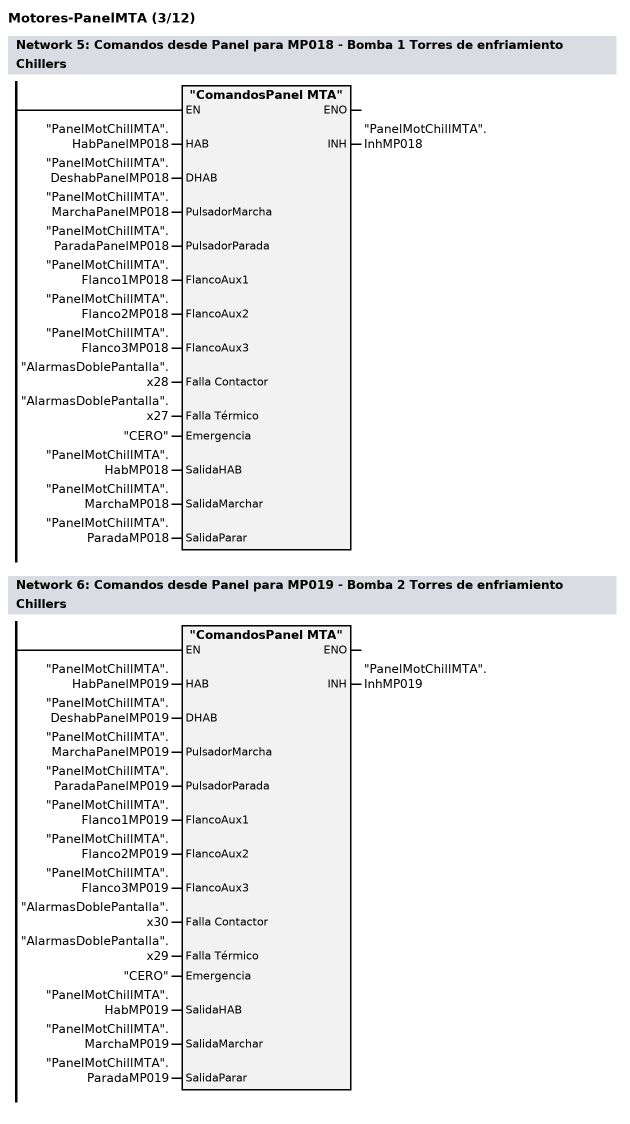
   RUNG wire#powerrail
      "ComandosPanel MTA"(HAB := "PanelMotChillMTA".HabPanelMP018, DHAB := "PanelMotChillMTA".DeshabPanelMP018, PulsadorMarcha := "PanelMotChillMTA".MarchaPanelMP018, PulsadorParada := "PanelMotChillMTA".ParadaPanelMP018, FlancoAux1 := "PanelMotChillMTA".Flanco1MP018, FlancoAux2 := "PanelMotChillMTA".Flanco2MP018, FlancoAux3 := "PanelMotChillMTA".Flanco3MP018, "Falla Contactor" := "AlarmasDoblePantalla".x28, "Falla Térmico" := "AlarmasDoblePantalla".x27, Emergencia := "CERO", SalidaHAB := "PanelMotChillMTA".HabMP018, SalidaMarchar := "PanelMotChillMTA".MarchaMP018, SalidaParar := "PanelMotChillMTA".ParadaMP018, INH => "PanelMotChillMTA".InhMP018)
   END_RUNG
   // the same network as SCL:
   "ComandosPanel MTA"(HAB := "PanelMotChillMTA".HabPanelMP018,
                       DHAB := "PanelMotChillMTA".DeshabPanelMP018,
                       PulsadorMarcha := "PanelMotChillMTA".MarchaPanelMP018,
                       PulsadorParada := "PanelMotChillMTA".ParadaPanelMP018,
                       FlancoAux1 := "PanelMotChillMTA".Flanco1MP018,
                       FlancoAux2 := "PanelMotChillMTA".Flanco2MP018,
                       FlancoAux3 := "PanelMotChillMTA".Flanco3MP018,
                       "Falla Contactor" := "AlarmasDoblePantalla".x28,
                       "Falla Térmico" := "AlarmasDoblePantalla".x27,
                       Emergencia := "CERO",
                       SalidaHAB := "PanelMotChillMTA".HabMP018,
                       SalidaMarchar := "PanelMotChillMTA".MarchaMP018,
                       SalidaParar := "PanelMotChillMTA".ParadaMP018,
                       INH => "PanelMotChillMTA".InhMP018);
END_REGION

REGION Network 6: Comandos desde Panel para MP019 - Bomba 2 Torres de enfriamiento Chillers
   RUNG wire#powerrail
      "ComandosPanel MTA"(HAB := "PanelMotChillMTA".HabPanelMP019, DHAB := "PanelMotChillMTA".DeshabPanelMP019, PulsadorMarcha := "PanelMotChillMTA".MarchaPanelMP019, PulsadorParada := "PanelMotChillMTA".ParadaPanelMP019, FlancoAux1 := "PanelMotChillMTA".Flanco1MP019, FlancoAux2 := "PanelMotChillMTA".Flanco2MP019, FlancoAux3 := "PanelMotChillMTA".Flanco3MP019, "Falla Contactor" := "AlarmasDoblePantalla".x30, "Falla Térmico" := "AlarmasDoblePantalla".x29, Emergencia := "CERO", SalidaHAB := "PanelMotChillMTA".HabMP019, SalidaMarchar := "PanelMotChillMTA".MarchaMP019, SalidaParar := "PanelMotChillMTA".ParadaMP019, INH => "PanelMotChillMTA".InhMP019)
   END_RUNG
   // the same network as SCL:
   "ComandosPanel MTA"(HAB := "PanelMotChillMTA".HabPanelMP019,
                       DHAB := "PanelMotChillMTA".DeshabPanelMP019,
                       PulsadorMarcha := "PanelMotChillMTA".MarchaPanelMP019,
                       PulsadorParada := "PanelMotChillMTA".ParadaPanelMP019,
                       FlancoAux1 := "PanelMotChillMTA".Flanco1MP019,
                       FlancoAux2 := "PanelMotChillMTA".Flanco2MP019,
                       FlancoAux3 := "PanelMotChillMTA".Flanco3MP019,
                       "Falla Contactor" := "AlarmasDoblePantalla".x30,
                       "Falla Térmico" := "AlarmasDoblePantalla".x29,
                       Emergencia := "CERO",
                       SalidaHAB := "PanelMotChillMTA".HabMP019,
                       SalidaMarchar := "PanelMotChillMTA".MarchaMP019,
                       SalidaParar := "PanelMotChillMTA".ParadaMP019,
                       INH => "PanelMotChillMTA".InhMP019);
END_REGION

REGION Network 7: Comandos desde Panel para MT007 - Bomba Soplado L1
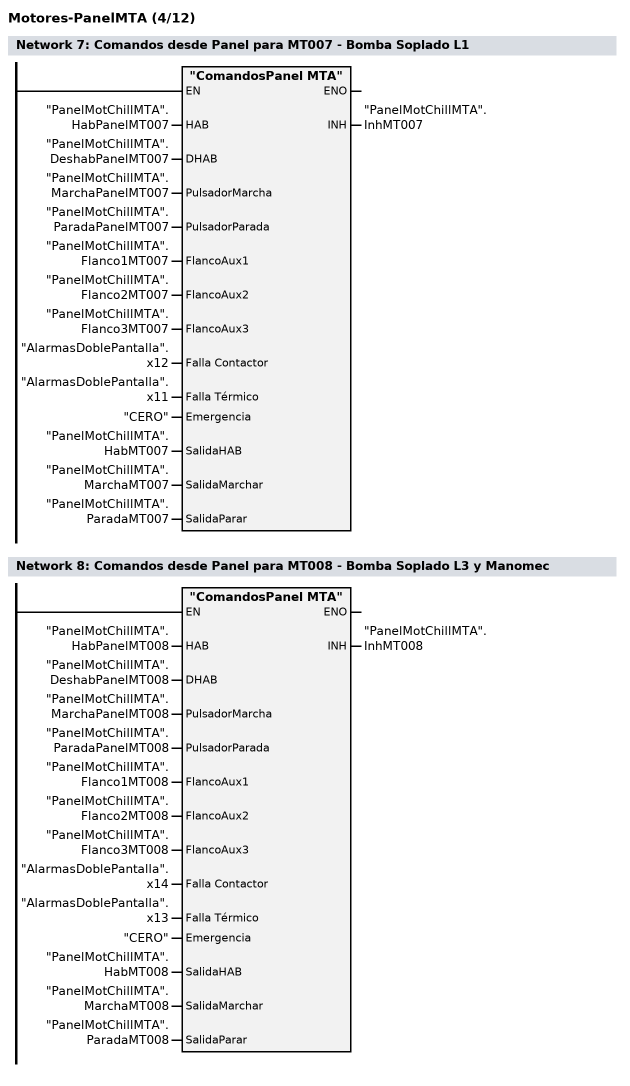
   RUNG wire#powerrail
      "ComandosPanel MTA"(HAB := "PanelMotChillMTA".HabPanelMT007, DHAB := "PanelMotChillMTA".DeshabPanelMT007, PulsadorMarcha := "PanelMotChillMTA".MarchaPanelMT007, PulsadorParada := "PanelMotChillMTA".ParadaPanelMT007, FlancoAux1 := "PanelMotChillMTA".Flanco1MT007, FlancoAux2 := "PanelMotChillMTA".Flanco2MT007, FlancoAux3 := "PanelMotChillMTA".Flanco3MT007, "Falla Contactor" := "AlarmasDoblePantalla".x12, "Falla Térmico" := "AlarmasDoblePantalla".x11, Emergencia := "CERO", INH => "PanelMotChillMTA".InhMT007, SalidaHAB := "PanelMotChillMTA".HabMT007, SalidaMarchar := "PanelMotChillMTA".MarchaMT007, SalidaParar := "PanelMotChillMTA".ParadaMT007)
   END_RUNG
   // the same network as SCL:
   "ComandosPanel MTA"(HAB := "PanelMotChillMTA".HabPanelMT007,
                       DHAB := "PanelMotChillMTA".DeshabPanelMT007,
                       PulsadorMarcha := "PanelMotChillMTA".MarchaPanelMT007,
                       PulsadorParada := "PanelMotChillMTA".ParadaPanelMT007,
                       FlancoAux1 := "PanelMotChillMTA".Flanco1MT007,
                       FlancoAux2 := "PanelMotChillMTA".Flanco2MT007,
                       FlancoAux3 := "PanelMotChillMTA".Flanco3MT007,
                       "Falla Contactor" := "AlarmasDoblePantalla".x12,
                       "Falla Térmico" := "AlarmasDoblePantalla".x11,
                       Emergencia := "CERO",
                       SalidaHAB := "PanelMotChillMTA".HabMT007,
                       SalidaMarchar := "PanelMotChillMTA".MarchaMT007,
                       SalidaParar := "PanelMotChillMTA".ParadaMT007,
                       INH => "PanelMotChillMTA".InhMT007);
END_REGION

REGION Network 8: Comandos desde Panel para MT008 - Bomba Soplado L3 y Manomec
   RUNG wire#powerrail
      "ComandosPanel MTA"(HAB := "PanelMotChillMTA".HabPanelMT008, DHAB := "PanelMotChillMTA".DeshabPanelMT008, PulsadorMarcha := "PanelMotChillMTA".MarchaPanelMT008, PulsadorParada := "PanelMotChillMTA".ParadaPanelMT008, FlancoAux1 := "PanelMotChillMTA".Flanco1MT008, FlancoAux2 := "PanelMotChillMTA".Flanco2MT008, FlancoAux3 := "PanelMotChillMTA".Flanco3MT008, "Falla Contactor" := "AlarmasDoblePantalla".x14, "Falla Térmico" := "AlarmasDoblePantalla".x13, Emergencia := "CERO", INH => "PanelMotChillMTA".InhMT008, SalidaHAB := "PanelMotChillMTA".HabMT008, SalidaMarchar := "PanelMotChillMTA".MarchaMT008, SalidaParar := "PanelMotChillMTA".ParadaMT008)
   END_RUNG
   // the same network as SCL:
   "ComandosPanel MTA"(HAB := "PanelMotChillMTA".HabPanelMT008,
                       DHAB := "PanelMotChillMTA".DeshabPanelMT008,
                       PulsadorMarcha := "PanelMotChillMTA".MarchaPanelMT008,
                       PulsadorParada := "PanelMotChillMTA".ParadaPanelMT008,
                       FlancoAux1 := "PanelMotChillMTA".Flanco1MT008,
                       FlancoAux2 := "PanelMotChillMTA".Flanco2MT008,
                       FlancoAux3 := "PanelMotChillMTA".Flanco3MT008,
                       "Falla Contactor" := "AlarmasDoblePantalla".x14,
                       "Falla Térmico" := "AlarmasDoblePantalla".x13,
                       Emergencia := "CERO",
                       SalidaHAB := "PanelMotChillMTA".HabMT008,
                       SalidaMarchar := "PanelMotChillMTA".MarchaMT008,
                       SalidaParar := "PanelMotChillMTA".ParadaMT008,
                       INH => "PanelMotChillMTA".InhMT008);
END_REGION

REGION Network 9: Comandos desde Panel para MT009 - Bomba Int. L3 y L5
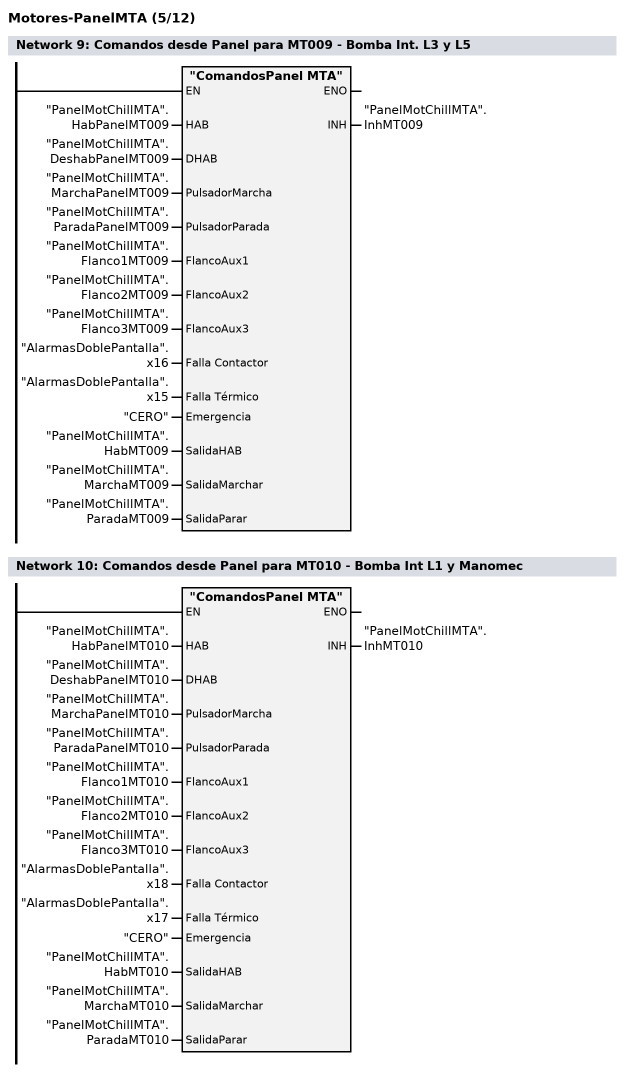
   RUNG wire#powerrail
      "ComandosPanel MTA"(HAB := "PanelMotChillMTA".HabPanelMT009, DHAB := "PanelMotChillMTA".DeshabPanelMT009, PulsadorMarcha := "PanelMotChillMTA".MarchaPanelMT009, PulsadorParada := "PanelMotChillMTA".ParadaPanelMT009, FlancoAux1 := "PanelMotChillMTA".Flanco1MT009, FlancoAux2 := "PanelMotChillMTA".Flanco2MT009, FlancoAux3 := "PanelMotChillMTA".Flanco3MT009, "Falla Contactor" := "AlarmasDoblePantalla".x16, "Falla Térmico" := "AlarmasDoblePantalla".x15, Emergencia := "CERO", INH => "PanelMotChillMTA".InhMT009, SalidaHAB := "PanelMotChillMTA".HabMT009, SalidaMarchar := "PanelMotChillMTA".MarchaMT009, SalidaParar := "PanelMotChillMTA".ParadaMT009)
   END_RUNG
   // the same network as SCL:
   "ComandosPanel MTA"(HAB := "PanelMotChillMTA".HabPanelMT009,
                       DHAB := "PanelMotChillMTA".DeshabPanelMT009,
                       PulsadorMarcha := "PanelMotChillMTA".MarchaPanelMT009,
                       PulsadorParada := "PanelMotChillMTA".ParadaPanelMT009,
                       FlancoAux1 := "PanelMotChillMTA".Flanco1MT009,
                       FlancoAux2 := "PanelMotChillMTA".Flanco2MT009,
                       FlancoAux3 := "PanelMotChillMTA".Flanco3MT009,
                       "Falla Contactor" := "AlarmasDoblePantalla".x16,
                       "Falla Térmico" := "AlarmasDoblePantalla".x15,
                       Emergencia := "CERO",
                       SalidaHAB := "PanelMotChillMTA".HabMT009,
                       SalidaMarchar := "PanelMotChillMTA".MarchaMT009,
                       SalidaParar := "PanelMotChillMTA".ParadaMT009,
                       INH => "PanelMotChillMTA".InhMT009);
END_REGION

REGION Network 10: Comandos desde Panel para MT010 - Bomba Int L1 y Manomec
   RUNG wire#powerrail
      "ComandosPanel MTA"(HAB := "PanelMotChillMTA".HabPanelMT010, DHAB := "PanelMotChillMTA".DeshabPanelMT010, PulsadorMarcha := "PanelMotChillMTA".MarchaPanelMT010, PulsadorParada := "PanelMotChillMTA".ParadaPanelMT010, FlancoAux1 := "PanelMotChillMTA".Flanco1MT010, FlancoAux2 := "PanelMotChillMTA".Flanco2MT010, FlancoAux3 := "PanelMotChillMTA".Flanco3MT010, "Falla Contactor" := "AlarmasDoblePantalla".x18, "Falla Térmico" := "AlarmasDoblePantalla".x17, Emergencia := "CERO", INH => "PanelMotChillMTA".InhMT010, SalidaHAB := "PanelMotChillMTA".HabMT010, SalidaMarchar := "PanelMotChillMTA".MarchaMT010, SalidaParar := "PanelMotChillMTA".ParadaMT010)
   END_RUNG
   // the same network as SCL:
   "ComandosPanel MTA"(HAB := "PanelMotChillMTA".HabPanelMT010,
                       DHAB := "PanelMotChillMTA".DeshabPanelMT010,
                       PulsadorMarcha := "PanelMotChillMTA".MarchaPanelMT010,
                       PulsadorParada := "PanelMotChillMTA".ParadaPanelMT010,
                       FlancoAux1 := "PanelMotChillMTA".Flanco1MT010,
                       FlancoAux2 := "PanelMotChillMTA".Flanco2MT010,
                       FlancoAux3 := "PanelMotChillMTA".Flanco3MT010,
                       "Falla Contactor" := "AlarmasDoblePantalla".x18,
                       "Falla Térmico" := "AlarmasDoblePantalla".x17,
                       Emergencia := "CERO",
                       SalidaHAB := "PanelMotChillMTA".HabMT010,
                       SalidaMarchar := "PanelMotChillMTA".MarchaMT010,
                       SalidaParar := "PanelMotChillMTA".ParadaMT010,
                       INH => "PanelMotChillMTA".InhMT010);
END_REGION

REGION Network 11: Comandos desde Panel para V001 - Ventilador 1 Torres de enfriamiento Chillers
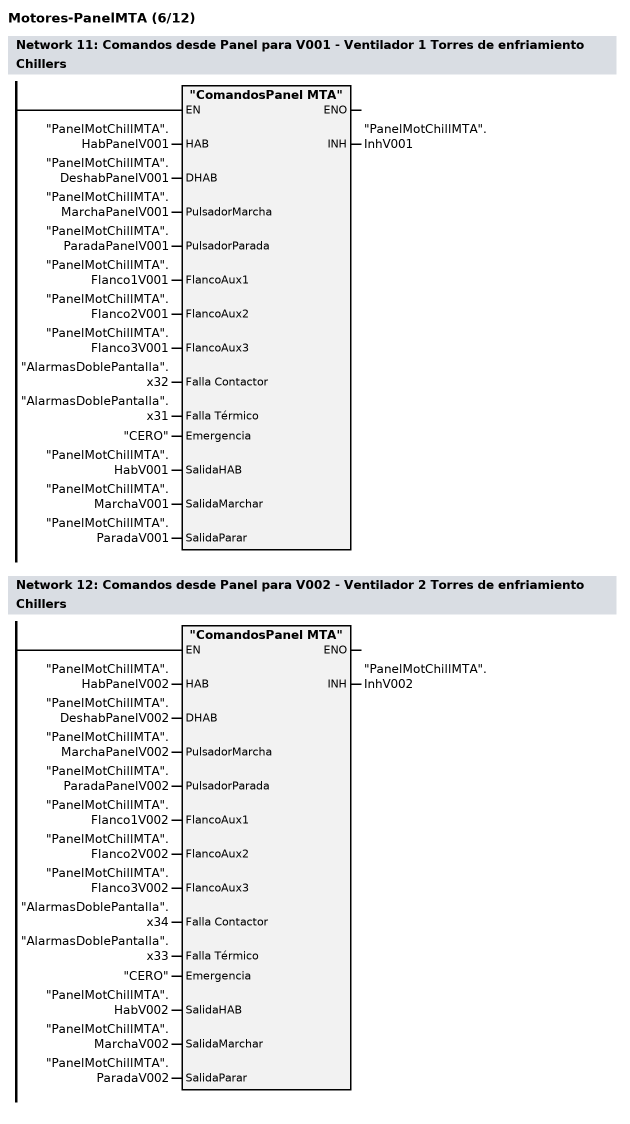
   RUNG wire#powerrail
      "ComandosPanel MTA"(HAB := "PanelMotChillMTA".HabPanelV001, DHAB := "PanelMotChillMTA".DeshabPanelV001, PulsadorMarcha := "PanelMotChillMTA".MarchaPanelV001, PulsadorParada := "PanelMotChillMTA".ParadaPanelV001, FlancoAux1 := "PanelMotChillMTA".Flanco1V001, FlancoAux2 := "PanelMotChillMTA".Flanco2V001, FlancoAux3 := "PanelMotChillMTA".Flanco3V001, "Falla Contactor" := "AlarmasDoblePantalla".x32, "Falla Térmico" := "AlarmasDoblePantalla".x31, Emergencia := "CERO", SalidaHAB := "PanelMotChillMTA".HabV001, SalidaMarchar := "PanelMotChillMTA".MarchaV001, SalidaParar := "PanelMotChillMTA".ParadaV001, INH => "PanelMotChillMTA".InhV001)
   END_RUNG
   // the same network as SCL:
   "ComandosPanel MTA"(HAB := "PanelMotChillMTA".HabPanelV001,
                       DHAB := "PanelMotChillMTA".DeshabPanelV001,
                       PulsadorMarcha := "PanelMotChillMTA".MarchaPanelV001,
                       PulsadorParada := "PanelMotChillMTA".ParadaPanelV001,
                       FlancoAux1 := "PanelMotChillMTA".Flanco1V001,
                       FlancoAux2 := "PanelMotChillMTA".Flanco2V001,
                       FlancoAux3 := "PanelMotChillMTA".Flanco3V001,
                       "Falla Contactor" := "AlarmasDoblePantalla".x32,
                       "Falla Térmico" := "AlarmasDoblePantalla".x31,
                       Emergencia := "CERO",
                       SalidaHAB := "PanelMotChillMTA".HabV001,
                       SalidaMarchar := "PanelMotChillMTA".MarchaV001,
                       SalidaParar := "PanelMotChillMTA".ParadaV001,
                       INH => "PanelMotChillMTA".InhV001);
END_REGION

REGION Network 12: Comandos desde Panel para V002 - Ventilador 2 Torres de enfriamiento Chillers
   RUNG wire#powerrail
      "ComandosPanel MTA"(HAB := "PanelMotChillMTA".HabPanelV002, DHAB := "PanelMotChillMTA".DeshabPanelV002, PulsadorMarcha := "PanelMotChillMTA".MarchaPanelV002, PulsadorParada := "PanelMotChillMTA".ParadaPanelV002, FlancoAux1 := "PanelMotChillMTA".Flanco1V002, FlancoAux2 := "PanelMotChillMTA".Flanco2V002, FlancoAux3 := "PanelMotChillMTA".Flanco3V002, "Falla Contactor" := "AlarmasDoblePantalla".x34, "Falla Térmico" := "AlarmasDoblePantalla".x33, Emergencia := "CERO", SalidaHAB := "PanelMotChillMTA".HabV002, SalidaMarchar := "PanelMotChillMTA".MarchaV002, SalidaParar := "PanelMotChillMTA".ParadaV002, INH => "PanelMotChillMTA".InhV002)
   END_RUNG
   // the same network as SCL:
   "ComandosPanel MTA"(HAB := "PanelMotChillMTA".HabPanelV002,
                       DHAB := "PanelMotChillMTA".DeshabPanelV002,
                       PulsadorMarcha := "PanelMotChillMTA".MarchaPanelV002,
                       PulsadorParada := "PanelMotChillMTA".ParadaPanelV002,
                       FlancoAux1 := "PanelMotChillMTA".Flanco1V002,
                       FlancoAux2 := "PanelMotChillMTA".Flanco2V002,
                       FlancoAux3 := "PanelMotChillMTA".Flanco3V002,
                       "Falla Contactor" := "AlarmasDoblePantalla".x34,
                       "Falla Térmico" := "AlarmasDoblePantalla".x33,
                       Emergencia := "CERO",
                       SalidaHAB := "PanelMotChillMTA".HabV002,
                       SalidaMarchar := "PanelMotChillMTA".MarchaV002,
                       SalidaParar := "PanelMotChillMTA".ParadaV002,
                       INH => "PanelMotChillMTA".InhV002);
END_REGION

REGION Network 13: Comandos desde Panel para V003 - Ventilador 3 Torres de enfriamiento Chillers
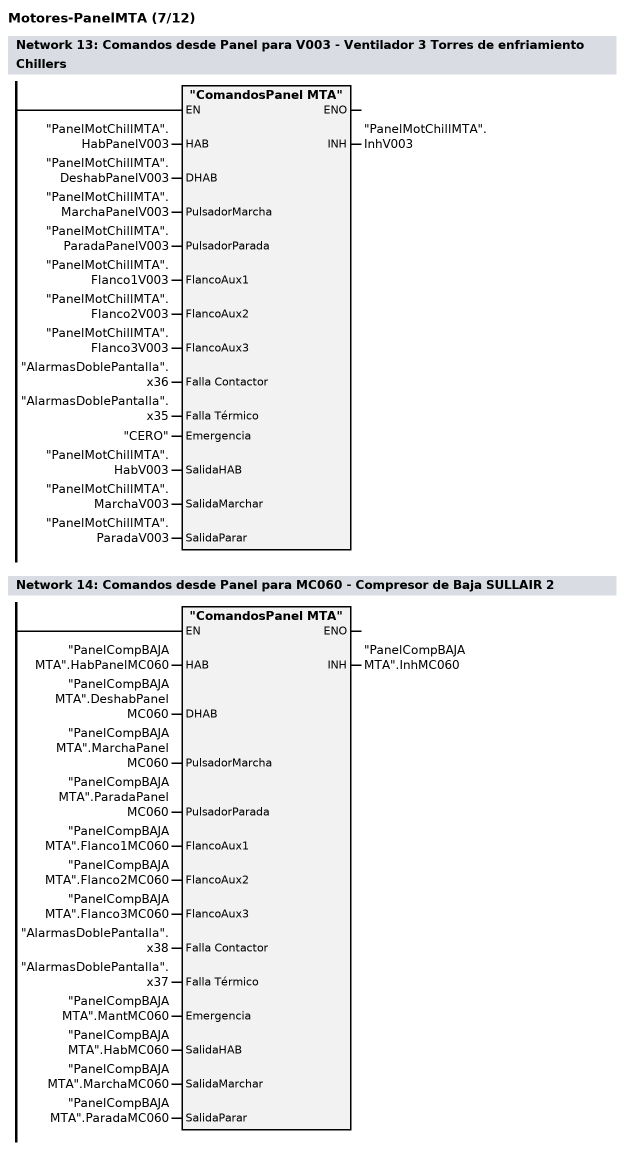
   RUNG wire#powerrail
      "ComandosPanel MTA"(HAB := "PanelMotChillMTA".HabPanelV003, DHAB := "PanelMotChillMTA".DeshabPanelV003, PulsadorMarcha := "PanelMotChillMTA".MarchaPanelV003, PulsadorParada := "PanelMotChillMTA".ParadaPanelV003, FlancoAux1 := "PanelMotChillMTA".Flanco1V003, FlancoAux2 := "PanelMotChillMTA".Flanco2V003, FlancoAux3 := "PanelMotChillMTA".Flanco3V003, "Falla Contactor" := "AlarmasDoblePantalla".x36, "Falla Térmico" := "AlarmasDoblePantalla".x35, Emergencia := "CERO", SalidaHAB := "PanelMotChillMTA".HabV003, SalidaMarchar := "PanelMotChillMTA".MarchaV003, SalidaParar := "PanelMotChillMTA".ParadaV003, INH => "PanelMotChillMTA".InhV003)
   END_RUNG
   // the same network as SCL:
   "ComandosPanel MTA"(HAB := "PanelMotChillMTA".HabPanelV003,
                       DHAB := "PanelMotChillMTA".DeshabPanelV003,
                       PulsadorMarcha := "PanelMotChillMTA".MarchaPanelV003,
                       PulsadorParada := "PanelMotChillMTA".ParadaPanelV003,
                       FlancoAux1 := "PanelMotChillMTA".Flanco1V003,
                       FlancoAux2 := "PanelMotChillMTA".Flanco2V003,
                       FlancoAux3 := "PanelMotChillMTA".Flanco3V003,
                       "Falla Contactor" := "AlarmasDoblePantalla".x36,
                       "Falla Térmico" := "AlarmasDoblePantalla".x35,
                       Emergencia := "CERO",
                       SalidaHAB := "PanelMotChillMTA".HabV003,
                       SalidaMarchar := "PanelMotChillMTA".MarchaV003,
                       SalidaParar := "PanelMotChillMTA".ParadaV003,
                       INH => "PanelMotChillMTA".InhV003);
END_REGION

REGION Network 14: Comandos desde Panel para MC060 - Compresor de Baja SULLAIR 2
   RUNG wire#powerrail
      "ComandosPanel MTA"(HAB := "PanelCompBAJA MTA".HabPanelMC060, DHAB := "PanelCompBAJA MTA".DeshabPanelMC060, PulsadorMarcha := "PanelCompBAJA MTA".MarchaPanelMC060, PulsadorParada := "PanelCompBAJA MTA".ParadaPanelMC060, FlancoAux1 := "PanelCompBAJA MTA".Flanco1MC060, FlancoAux2 := "PanelCompBAJA MTA".Flanco2MC060, FlancoAux3 := "PanelCompBAJA MTA".Flanco3MC060, "Falla Contactor" := "AlarmasDoblePantalla".x38, "Falla Térmico" := "AlarmasDoblePantalla".x37, Emergencia := "PanelCompBAJA MTA".MantMC060, INH => "PanelCompBAJA MTA".InhMC060, SalidaHAB := "PanelCompBAJA MTA".HabMC060, SalidaMarchar := "PanelCompBAJA MTA".MarchaMC060, SalidaParar := "PanelCompBAJA MTA".ParadaMC060)
   END_RUNG
   // the same network as SCL:
   "ComandosPanel MTA"(HAB := "PanelCompBAJA MTA".HabPanelMC060,
                       DHAB := "PanelCompBAJA MTA".DeshabPanelMC060,
                       PulsadorMarcha := "PanelCompBAJA MTA".MarchaPanelMC060,
                       PulsadorParada := "PanelCompBAJA MTA".ParadaPanelMC060,
                       FlancoAux1 := "PanelCompBAJA MTA".Flanco1MC060,
                       FlancoAux2 := "PanelCompBAJA MTA".Flanco2MC060,
                       FlancoAux3 := "PanelCompBAJA MTA".Flanco3MC060,
                       "Falla Contactor" := "AlarmasDoblePantalla".x38,
                       "Falla Térmico" := "AlarmasDoblePantalla".x37,
                       Emergencia := "PanelCompBAJA MTA".MantMC060,
                       SalidaHAB := "PanelCompBAJA MTA".HabMC060,
                       SalidaMarchar := "PanelCompBAJA MTA".MarchaMC060,
                       SalidaParar := "PanelCompBAJA MTA".ParadaMC060,
                       INH => "PanelCompBAJA MTA".InhMC060);
END_REGION

REGION Network 15: Comandos desde Panel para MC061 - Compresor de Baja SULLAIR 1
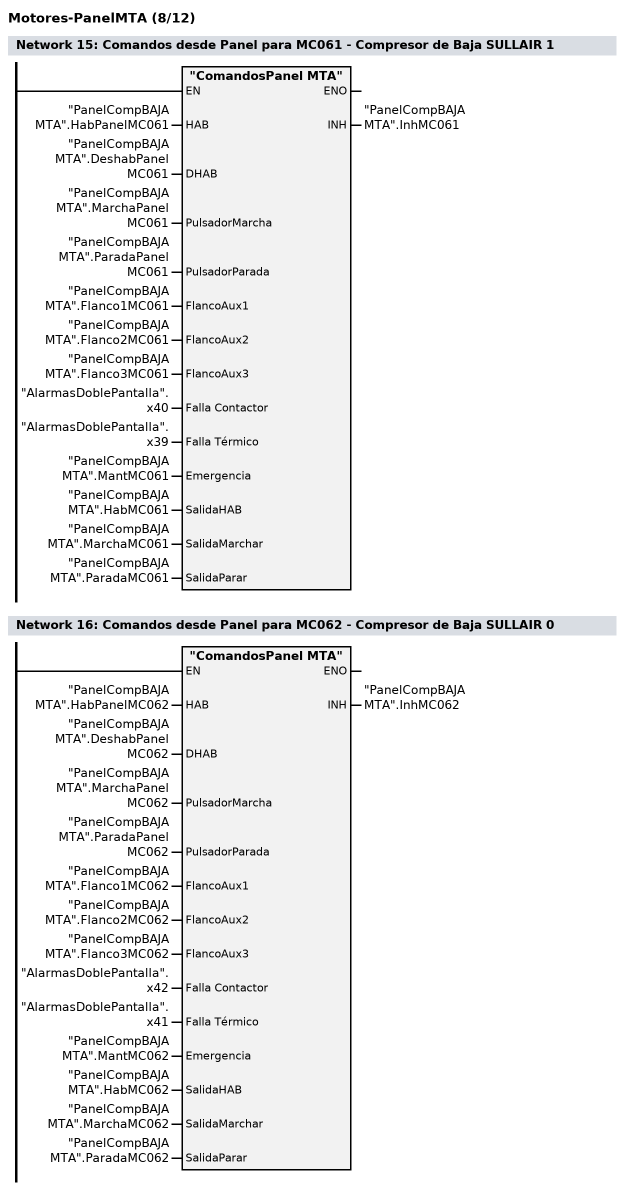
   RUNG wire#powerrail
      "ComandosPanel MTA"(HAB := "PanelCompBAJA MTA".HabPanelMC061, DHAB := "PanelCompBAJA MTA".DeshabPanelMC061, PulsadorMarcha := "PanelCompBAJA MTA".MarchaPanelMC061, PulsadorParada := "PanelCompBAJA MTA".ParadaPanelMC061, FlancoAux1 := "PanelCompBAJA MTA".Flanco1MC061, FlancoAux2 := "PanelCompBAJA MTA".Flanco2MC061, FlancoAux3 := "PanelCompBAJA MTA".Flanco3MC061, "Falla Contactor" := "AlarmasDoblePantalla".x40, "Falla Térmico" := "AlarmasDoblePantalla".x39, Emergencia := "PanelCompBAJA MTA".MantMC061, INH => "PanelCompBAJA MTA".InhMC061, SalidaHAB := "PanelCompBAJA MTA".HabMC061, SalidaMarchar := "PanelCompBAJA MTA".MarchaMC061, SalidaParar := "PanelCompBAJA MTA".ParadaMC061)
   END_RUNG
   // the same network as SCL:
   "ComandosPanel MTA"(HAB := "PanelCompBAJA MTA".HabPanelMC061,
                       DHAB := "PanelCompBAJA MTA".DeshabPanelMC061,
                       PulsadorMarcha := "PanelCompBAJA MTA".MarchaPanelMC061,
                       PulsadorParada := "PanelCompBAJA MTA".ParadaPanelMC061,
                       FlancoAux1 := "PanelCompBAJA MTA".Flanco1MC061,
                       FlancoAux2 := "PanelCompBAJA MTA".Flanco2MC061,
                       FlancoAux3 := "PanelCompBAJA MTA".Flanco3MC061,
                       "Falla Contactor" := "AlarmasDoblePantalla".x40,
                       "Falla Térmico" := "AlarmasDoblePantalla".x39,
                       Emergencia := "PanelCompBAJA MTA".MantMC061,
                       SalidaHAB := "PanelCompBAJA MTA".HabMC061,
                       SalidaMarchar := "PanelCompBAJA MTA".MarchaMC061,
                       SalidaParar := "PanelCompBAJA MTA".ParadaMC061,
                       INH => "PanelCompBAJA MTA".InhMC061);
END_REGION

REGION Network 16: Comandos desde Panel para MC062 - Compresor de Baja SULLAIR 0
   RUNG wire#powerrail
      "ComandosPanel MTA"(HAB := "PanelCompBAJA MTA".HabPanelMC062, DHAB := "PanelCompBAJA MTA".DeshabPanelMC062, PulsadorMarcha := "PanelCompBAJA MTA".MarchaPanelMC062, PulsadorParada := "PanelCompBAJA MTA".ParadaPanelMC062, FlancoAux1 := "PanelCompBAJA MTA".Flanco1MC062, FlancoAux2 := "PanelCompBAJA MTA".Flanco2MC062, FlancoAux3 := "PanelCompBAJA MTA".Flanco3MC062, "Falla Contactor" := "AlarmasDoblePantalla".x42, "Falla Térmico" := "AlarmasDoblePantalla".x41, Emergencia := "PanelCompBAJA MTA".MantMC062, INH => "PanelCompBAJA MTA".InhMC062, SalidaHAB := "PanelCompBAJA MTA".HabMC062, SalidaMarchar := "PanelCompBAJA MTA".MarchaMC062, SalidaParar := "PanelCompBAJA MTA".ParadaMC062)
   END_RUNG
   // the same network as SCL:
   "ComandosPanel MTA"(HAB := "PanelCompBAJA MTA".HabPanelMC062,
                       DHAB := "PanelCompBAJA MTA".DeshabPanelMC062,
                       PulsadorMarcha := "PanelCompBAJA MTA".MarchaPanelMC062,
                       PulsadorParada := "PanelCompBAJA MTA".ParadaPanelMC062,
                       FlancoAux1 := "PanelCompBAJA MTA".Flanco1MC062,
                       FlancoAux2 := "PanelCompBAJA MTA".Flanco2MC062,
                       FlancoAux3 := "PanelCompBAJA MTA".Flanco3MC062,
                       "Falla Contactor" := "AlarmasDoblePantalla".x42,
                       "Falla Térmico" := "AlarmasDoblePantalla".x41,
                       Emergencia := "PanelCompBAJA MTA".MantMC062,
                       SalidaHAB := "PanelCompBAJA MTA".HabMC062,
                       SalidaMarchar := "PanelCompBAJA MTA".MarchaMC062,
                       SalidaParar := "PanelCompBAJA MTA".ParadaMC062,
                       INH => "PanelCompBAJA MTA".InhMC062);
END_REGION

REGION Network 17: Comandos desde Panel para MC063 - Compresor de Baja ATLAS 3
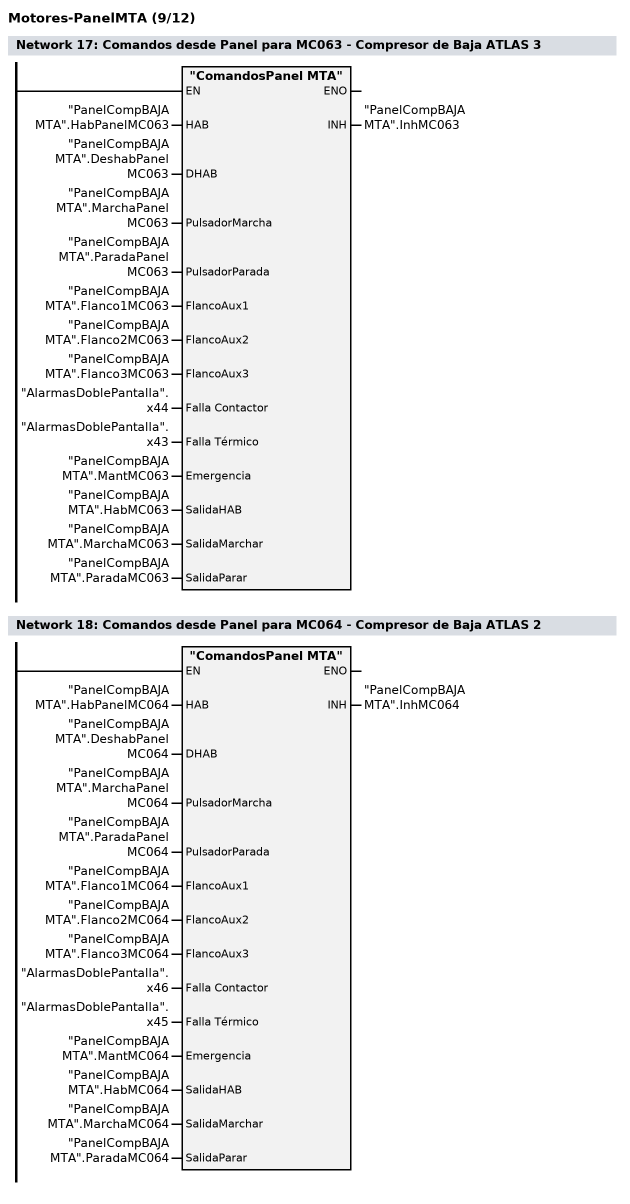
   RUNG wire#powerrail
      "ComandosPanel MTA"(HAB := "PanelCompBAJA MTA".HabPanelMC063, DHAB := "PanelCompBAJA MTA".DeshabPanelMC063, PulsadorMarcha := "PanelCompBAJA MTA".MarchaPanelMC063, PulsadorParada := "PanelCompBAJA MTA".ParadaPanelMC063, FlancoAux1 := "PanelCompBAJA MTA".Flanco1MC063, FlancoAux2 := "PanelCompBAJA MTA".Flanco2MC063, FlancoAux3 := "PanelCompBAJA MTA".Flanco3MC063, "Falla Contactor" := "AlarmasDoblePantalla".x44, "Falla Térmico" := "AlarmasDoblePantalla".x43, Emergencia := "PanelCompBAJA MTA".MantMC063, INH => "PanelCompBAJA MTA".InhMC063, SalidaHAB := "PanelCompBAJA MTA".HabMC063, SalidaMarchar := "PanelCompBAJA MTA".MarchaMC063, SalidaParar := "PanelCompBAJA MTA".ParadaMC063)
   END_RUNG
   // the same network as SCL:
   "ComandosPanel MTA"(HAB := "PanelCompBAJA MTA".HabPanelMC063,
                       DHAB := "PanelCompBAJA MTA".DeshabPanelMC063,
                       PulsadorMarcha := "PanelCompBAJA MTA".MarchaPanelMC063,
                       PulsadorParada := "PanelCompBAJA MTA".ParadaPanelMC063,
                       FlancoAux1 := "PanelCompBAJA MTA".Flanco1MC063,
                       FlancoAux2 := "PanelCompBAJA MTA".Flanco2MC063,
                       FlancoAux3 := "PanelCompBAJA MTA".Flanco3MC063,
                       "Falla Contactor" := "AlarmasDoblePantalla".x44,
                       "Falla Térmico" := "AlarmasDoblePantalla".x43,
                       Emergencia := "PanelCompBAJA MTA".MantMC063,
                       SalidaHAB := "PanelCompBAJA MTA".HabMC063,
                       SalidaMarchar := "PanelCompBAJA MTA".MarchaMC063,
                       SalidaParar := "PanelCompBAJA MTA".ParadaMC063,
                       INH => "PanelCompBAJA MTA".InhMC063);
END_REGION

REGION Network 18: Comandos desde Panel para MC064 - Compresor de Baja ATLAS 2
   RUNG wire#powerrail
      "ComandosPanel MTA"(HAB := "PanelCompBAJA MTA".HabPanelMC064, DHAB := "PanelCompBAJA MTA".DeshabPanelMC064, PulsadorMarcha := "PanelCompBAJA MTA".MarchaPanelMC064, PulsadorParada := "PanelCompBAJA MTA".ParadaPanelMC064, FlancoAux1 := "PanelCompBAJA MTA".Flanco1MC064, FlancoAux2 := "PanelCompBAJA MTA".Flanco2MC064, FlancoAux3 := "PanelCompBAJA MTA".Flanco3MC064, "Falla Contactor" := "AlarmasDoblePantalla".x46, "Falla Térmico" := "AlarmasDoblePantalla".x45, Emergencia := "PanelCompBAJA MTA".MantMC064, INH => "PanelCompBAJA MTA".InhMC064, SalidaHAB := "PanelCompBAJA MTA".HabMC064, SalidaMarchar := "PanelCompBAJA MTA".MarchaMC064, SalidaParar := "PanelCompBAJA MTA".ParadaMC064)
   END_RUNG
   // the same network as SCL:
   "ComandosPanel MTA"(HAB := "PanelCompBAJA MTA".HabPanelMC064,
                       DHAB := "PanelCompBAJA MTA".DeshabPanelMC064,
                       PulsadorMarcha := "PanelCompBAJA MTA".MarchaPanelMC064,
                       PulsadorParada := "PanelCompBAJA MTA".ParadaPanelMC064,
                       FlancoAux1 := "PanelCompBAJA MTA".Flanco1MC064,
                       FlancoAux2 := "PanelCompBAJA MTA".Flanco2MC064,
                       FlancoAux3 := "PanelCompBAJA MTA".Flanco3MC064,
                       "Falla Contactor" := "AlarmasDoblePantalla".x46,
                       "Falla Térmico" := "AlarmasDoblePantalla".x45,
                       Emergencia := "PanelCompBAJA MTA".MantMC064,
                       SalidaHAB := "PanelCompBAJA MTA".HabMC064,
                       SalidaMarchar := "PanelCompBAJA MTA".MarchaMC064,
                       SalidaParar := "PanelCompBAJA MTA".ParadaMC064,
                       INH => "PanelCompBAJA MTA".InhMC064);
END_REGION

REGION Network 19: Comandos desde Panel para MS050 - Secador de Alta ABC1
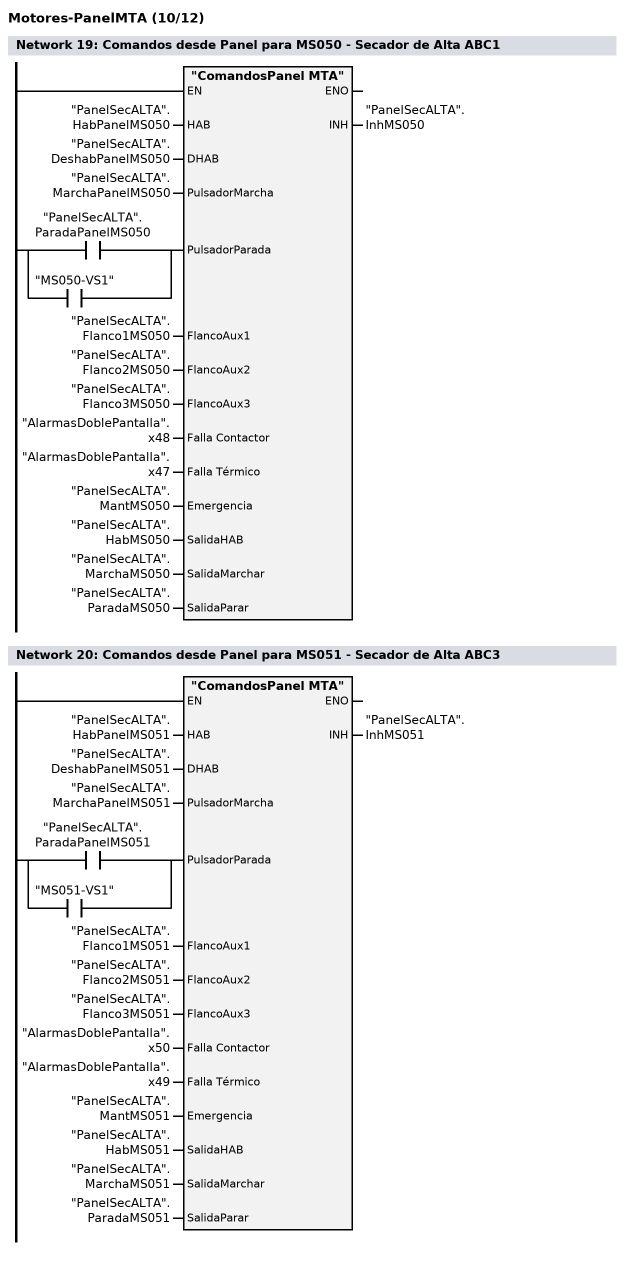
   RUNG wire#powerrail
      "ComandosPanel MTA"(HAB := "PanelSecALTA".HabPanelMS050, DHAB := "PanelSecALTA".DeshabPanelMS050, PulsadorMarcha := "PanelSecALTA".MarchaPanelMS050, PulsadorParada := wire#w1, FlancoAux1 := "PanelSecALTA".Flanco1MS050, FlancoAux2 := "PanelSecALTA".Flanco2MS050, FlancoAux3 := "PanelSecALTA".Flanco3MS050, "Falla Contactor" := "AlarmasDoblePantalla".x48, "Falla Térmico" := "AlarmasDoblePantalla".x47, Emergencia := "PanelSecALTA".MantMS050, INH => "PanelSecALTA".InhMS050, SalidaHAB := "PanelSecALTA".HabMS050, SalidaMarchar := "PanelSecALTA".MarchaMS050, SalidaParar := "PanelSecALTA".ParadaMS050)
   END_RUNG
   RUNG wire#powerrail
      Contact( "PanelSecALTA".ParadaPanelMS050 )
   END_RUNG wire#w1
   RUNG wire#powerrail
      Contact( "MS050-VS1" )
   END_RUNG wire#w1
   // the same network as SCL:
   "ComandosPanel MTA"(HAB := "PanelSecALTA".HabPanelMS050,
                       DHAB := "PanelSecALTA".DeshabPanelMS050,
                       PulsadorMarcha := "PanelSecALTA".MarchaPanelMS050,
                       PulsadorParada := "PanelSecALTA".ParadaPanelMS050 OR "MS050-VS1",
                       FlancoAux1 := "PanelSecALTA".Flanco1MS050,
                       FlancoAux2 := "PanelSecALTA".Flanco2MS050,
                       FlancoAux3 := "PanelSecALTA".Flanco3MS050,
                       "Falla Contactor" := "AlarmasDoblePantalla".x48,
                       "Falla Térmico" := "AlarmasDoblePantalla".x47,
                       Emergencia := "PanelSecALTA".MantMS050,
                       SalidaHAB := "PanelSecALTA".HabMS050,
                       SalidaMarchar := "PanelSecALTA".MarchaMS050,
                       SalidaParar := "PanelSecALTA".ParadaMS050,
                       INH => "PanelSecALTA".InhMS050);
END_REGION

REGION Network 20: Comandos desde Panel para MS051 - Secador de Alta ABC3
   RUNG wire#powerrail
      "ComandosPanel MTA"(HAB := "PanelSecALTA".HabPanelMS051, DHAB := "PanelSecALTA".DeshabPanelMS051, PulsadorMarcha := "PanelSecALTA".MarchaPanelMS051, PulsadorParada := wire#w1, FlancoAux1 := "PanelSecALTA".Flanco1MS051, FlancoAux2 := "PanelSecALTA".Flanco2MS051, FlancoAux3 := "PanelSecALTA".Flanco3MS051, "Falla Contactor" := "AlarmasDoblePantalla".x50, "Falla Térmico" := "AlarmasDoblePantalla".x49, Emergencia := "PanelSecALTA".MantMS051, INH => "PanelSecALTA".InhMS051, SalidaHAB := "PanelSecALTA".HabMS051, SalidaMarchar := "PanelSecALTA".MarchaMS051, SalidaParar := "PanelSecALTA".ParadaMS051)
   END_RUNG
   RUNG wire#powerrail
      Contact( "PanelSecALTA".ParadaPanelMS051 )
   END_RUNG wire#w1
   RUNG wire#powerrail
      Contact( "MS051-VS1" )
   END_RUNG wire#w1
   // the same network as SCL:
   "ComandosPanel MTA"(HAB := "PanelSecALTA".HabPanelMS051,
                       DHAB := "PanelSecALTA".DeshabPanelMS051,
                       PulsadorMarcha := "PanelSecALTA".MarchaPanelMS051,
                       PulsadorParada := "PanelSecALTA".ParadaPanelMS051 OR "MS051-VS1",
                       FlancoAux1 := "PanelSecALTA".Flanco1MS051,
                       FlancoAux2 := "PanelSecALTA".Flanco2MS051,
                       FlancoAux3 := "PanelSecALTA".Flanco3MS051,
                       "Falla Contactor" := "AlarmasDoblePantalla".x50,
                       "Falla Térmico" := "AlarmasDoblePantalla".x49,
                       Emergencia := "PanelSecALTA".MantMS051,
                       SalidaHAB := "PanelSecALTA".HabMS051,
                       SalidaMarchar := "PanelSecALTA".MarchaMS051,
                       SalidaParar := "PanelSecALTA".ParadaMS051,
                       INH => "PanelSecALTA".InhMS051);
END_REGION

REGION Network 21: Comandos desde Panel para MS052 - Secador de Alta ABC2
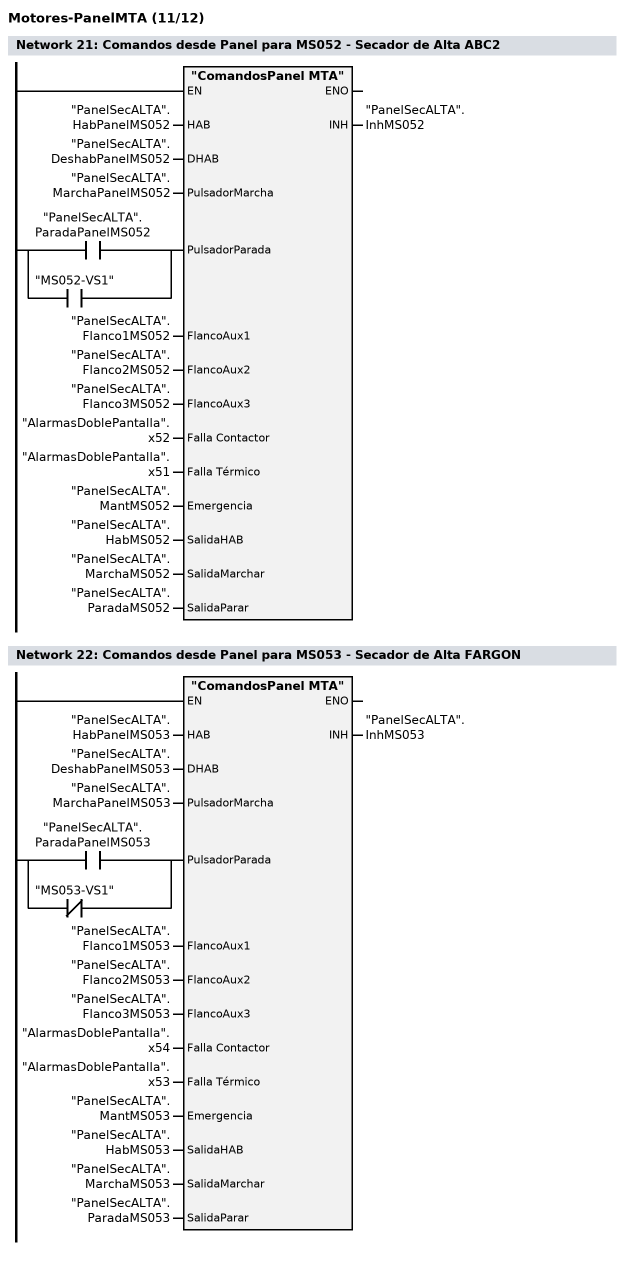
   RUNG wire#powerrail
      "ComandosPanel MTA"(HAB := "PanelSecALTA".HabPanelMS052, DHAB := "PanelSecALTA".DeshabPanelMS052, PulsadorMarcha := "PanelSecALTA".MarchaPanelMS052, PulsadorParada := wire#w1, FlancoAux1 := "PanelSecALTA".Flanco1MS052, FlancoAux2 := "PanelSecALTA".Flanco2MS052, FlancoAux3 := "PanelSecALTA".Flanco3MS052, "Falla Contactor" := "AlarmasDoblePantalla".x52, "Falla Térmico" := "AlarmasDoblePantalla".x51, Emergencia := "PanelSecALTA".MantMS052, INH => "PanelSecALTA".InhMS052, SalidaHAB := "PanelSecALTA".HabMS052, SalidaMarchar := "PanelSecALTA".MarchaMS052, SalidaParar := "PanelSecALTA".ParadaMS052)
   END_RUNG
   RUNG wire#powerrail
      Contact( "PanelSecALTA".ParadaPanelMS052 )
   END_RUNG wire#w1
   RUNG wire#powerrail
      Contact( "MS052-VS1" )
   END_RUNG wire#w1
   // the same network as SCL:
   "ComandosPanel MTA"(HAB := "PanelSecALTA".HabPanelMS052,
                       DHAB := "PanelSecALTA".DeshabPanelMS052,
                       PulsadorMarcha := "PanelSecALTA".MarchaPanelMS052,
                       PulsadorParada := "PanelSecALTA".ParadaPanelMS052 OR "MS052-VS1",
                       FlancoAux1 := "PanelSecALTA".Flanco1MS052,
                       FlancoAux2 := "PanelSecALTA".Flanco2MS052,
                       FlancoAux3 := "PanelSecALTA".Flanco3MS052,
                       "Falla Contactor" := "AlarmasDoblePantalla".x52,
                       "Falla Térmico" := "AlarmasDoblePantalla".x51,
                       Emergencia := "PanelSecALTA".MantMS052,
                       SalidaHAB := "PanelSecALTA".HabMS052,
                       SalidaMarchar := "PanelSecALTA".MarchaMS052,
                       SalidaParar := "PanelSecALTA".ParadaMS052,
                       INH => "PanelSecALTA".InhMS052);
END_REGION

REGION Network 22: Comandos desde Panel para MS053 - Secador de Alta FARGON
   RUNG wire#powerrail
      "ComandosPanel MTA"(HAB := "PanelSecALTA".HabPanelMS053, DHAB := "PanelSecALTA".DeshabPanelMS053, PulsadorMarcha := "PanelSecALTA".MarchaPanelMS053, PulsadorParada := wire#w1, FlancoAux1 := "PanelSecALTA".Flanco1MS053, FlancoAux2 := "PanelSecALTA".Flanco2MS053, FlancoAux3 := "PanelSecALTA".Flanco3MS053, "Falla Contactor" := "AlarmasDoblePantalla".x54, "Falla Térmico" := "AlarmasDoblePantalla".x53, Emergencia := "PanelSecALTA".MantMS053, INH => "PanelSecALTA".InhMS053, SalidaHAB := "PanelSecALTA".HabMS053, SalidaMarchar := "PanelSecALTA".MarchaMS053, SalidaParar := "PanelSecALTA".ParadaMS053)
   END_RUNG
   RUNG wire#powerrail
      Contact( "PanelSecALTA".ParadaPanelMS053 )
   END_RUNG wire#w1
   RUNG wire#powerrail
      I_Contact( "MS053-VS1" )
   END_RUNG wire#w1
   // the same network as SCL:
   "ComandosPanel MTA"(HAB := "PanelSecALTA".HabPanelMS053,
                       DHAB := "PanelSecALTA".DeshabPanelMS053,
                       PulsadorMarcha := "PanelSecALTA".MarchaPanelMS053,
                       PulsadorParada := "PanelSecALTA".ParadaPanelMS053 OR NOT "MS053-VS1",
                       FlancoAux1 := "PanelSecALTA".Flanco1MS053,
                       FlancoAux2 := "PanelSecALTA".Flanco2MS053,
                       FlancoAux3 := "PanelSecALTA".Flanco3MS053,
                       "Falla Contactor" := "AlarmasDoblePantalla".x54,
                       "Falla Térmico" := "AlarmasDoblePantalla".x53,
                       Emergencia := "PanelSecALTA".MantMS053,
                       SalidaHAB := "PanelSecALTA".HabMS053,
                       SalidaMarchar := "PanelSecALTA".MarchaMS053,
                       SalidaParar := "PanelSecALTA".ParadaMS053,
                       INH => "PanelSecALTA".InhMS053);
END_REGION

REGION Network 23: Comandos desde Panel para MS054 - Secador de Baja SULLAIR 1